
discrete alarms
   1: '', class Errors, trigger "Alarm0Pack16B_Alarmas_word" bit 0
   2: '', class Errors, trigger "Alarm0Pack16B_Alarmas_word" bit 1
   3: '', class Errors, trigger "Alarm0Pack16B_Alarmas_word" bit 2
   4: '', class Errors, trigger "Alarm0Pack16B_Alarmas_word" bit 3
   5: '', class Errors, trigger "Alarm0Pack16B_Alarmas_word" bit 4
   6: '', class Errors, trigger "Alarm0Pack16B_Alarmas_word" bit 5
   7: '', class Errors, trigger "Alarm0Pack16B_Alarmas_word" bit 6
   8: '', class Errors, trigger "Alarm0Pack16B_Alarmas_word" bit 7
   9: '', class Errors, trigger "Alarm0Pack16B_Alarmas_word" bit 8
   10: '', class Errors, trigger "Alarm0Pack16B_Alarmas_word" bit 9
   11: '', class Errors, trigger "Alarm0Pack16B_Alarmas_word" bit 10
   12: '', class Errors, trigger "Alarm0Pack16B_Alarmas_word" bit 11
   13: '', class Errors, trigger "Alarm0Pack16B_Alarmas_word" bit 12
   14: '', class Errors, trigger "Alarm0Pack16B_Alarmas_word" bit 13
   15: '', class Errors, trigger "Alarm0Pack16B_Alarmas_word" bit 14
   16: '', class Errors, trigger "Alarm0Pack16B_Alarmas_word" bit 15
   17: 'PeakDisplayPreAlarmHI', class Errors, trigger "Alarm1Pack16B_Alarmas_word" bit 0
   18: 'PeakDisplayAlarmHI', class Errors, trigger "Alarm1Pack16B_Alarmas_word" bit 1
   19: 'PeakDisplayPreAlarmLOW', class Errors, trigger "Alarm1Pack16B_Alarmas_word" bit 2
   20: 'PeakDisplayAlarmLOW', class Errors, trigger "Alarm1Pack16B_Alarmas_word" bit 3
   21: 'PlateauDisplayPreAlarmHI', class Errors, trigger "Alarm1Pack16B_Alarmas_word" bit 4
   22: 'PlateauDisplayAlarmHI', class Errors, trigger "Alarm1Pack16B_Alarmas_word" bit 5
   23: 'PlateauDisplayPreAlarmLOW', class Errors, trigger "Alarm1Pack16B_Alarmas_word" bit 6
   24: 'PlateaukDisplayAlarmLOW', class Errors, trigger "Alarm1Pack16B_Alarmas_word" bit 7
   25: 'PeepDisplayPreAlarmHI', class Errors, trigger "Alarm1Pack16B_Alarmas_word" bit 8
   26: 'PeepDisplayAlarmHI', class Errors, trigger "Alarm1Pack16B_Alarmas_word" bit 9
   27: 'PeepDisplayPreAlarmLOW', class Errors, trigger "Alarm1Pack16B_Alarmas_word" bit 10
   28: 'PeepDisplayAlarmLOW', class Errors, trigger "Alarm1Pack16B_Alarmas_word" bit 11
   29: 'FrequenciaDisplayPreAlarm / FrequencyDisplayPreAlarm', class Errors, trigger "Alarm1Pack16B_Alarmas_word" bit 12
   30: 'FrequenciaDisplayAlarmHI / FrequencyDisplayAlarmHI', class Errors, trigger "Alarm1Pack16B_Alarmas_word" bit 13
   31: 'FrequenciaDisplayPreAlarmLOW / FrequencyDisplayPreAlarmLOW', class Errors, trigger "Alarm1Pack16B_Alarmas_word" bit 14
   32: 'FrequenciaDisplayAlarmLOW / FrequencyDisplayAlarmLOW', class Errors, trigger "Alarm1Pack16B_Alarmas_word" bit 15
   33: 'TidalVolumeDisplayPreAlarm', class Errors, trigger "Alarm2Pack16B_Alarmas_word" bit 0
   34: 'TidalVolumeDisplayAlarmHI', class Errors, trigger "Alarm2Pack16B_Alarmas_word" bit 1
   35: 'TidalVolumeDisplayPreAlarmLOW', class Errors, trigger "Alarm2Pack16B_Alarmas_word" bit 2
   36: 'TidalVolumeDisplayAlarmLOW', class Errors, trigger "Alarm2Pack16B_Alarmas_word" bit 3
   37: 'MinuteVolumeDisplayPreAlarm', class Errors, trigger "Alarm2Pack16B_Alarmas_word" bit 4
   38: 'MinuteVolumeDisplayAlarmHI', class Errors, trigger "Alarm2Pack16B_Alarmas_word" bit 5
   39: 'MinuteVolumeDisplayPreAlarmLOW', class Errors, trigger "Alarm2Pack16B_Alarmas_word" bit 6
   40: 'MinuteVolumeDisplayAlarmLOW', class Errors, trigger "Alarm2Pack16B_Alarmas_word" bit 7
   41: 'TriggerDisplayPreAlarm', class Errors, trigger "Alarm2Pack16B_Alarmas_word" bit 8
   42: 'TriggerVolumeDisplayAlarmHI', class Errors, trigger "Alarm2Pack16B_Alarmas_word" bit 9
   43: 'TriggerVolumeDisplayPreAlarmLOW', class Errors, trigger "Alarm2Pack16B_Alarmas_word" bit 10
   44: 'TriggerVolumeDisplayAlarmLOW', class Errors, trigger "Alarm2Pack16B_Alarmas_word" bit 11
   45: 'BatteryDisplayPreAlarmHI', class Errors, trigger "Alarm2Pack16B_Alarmas_word" bit 12
   46: 'BatteryDisplayAlarmHI', class Errors, trigger "Alarm2Pack16B_Alarmas_word" bit 13
   47: 'BatteryDisplayPreAlarmLOW', class Errors, trigger "Alarm2Pack16B_Alarmas_word" bit 14
   48: 'BatteryDisplayAlarmLOW', class Errors, trigger "Alarm2Pack16B_Alarmas_word" bit 15
   49: '', class Errors, trigger "Alarm3Pack16B_Alarmas_word" bit 0
   50: '', class Errors, trigger "Alarm3Pack16B_Alarmas_word" bit 1
   51: '', class Errors, trigger "Alarm3Pack16B_Alarmas_word" bit 2
   52: '', class Errors, trigger "Alarm3Pack16B_Alarmas_word" bit 3
   53: '', class Errors, trigger "Alarm3Pack16B_Alarmas_word" bit 4
   54: '', class Errors, trigger "Alarm3Pack16B_Alarmas_word" bit 5
   55: '', class Errors, trigger "Alarm3Pack16B_Alarmas_word" bit 6
   56: '', class Errors, trigger "Alarm3Pack16B_Alarmas_word" bit 7
   57: '', class Errors, trigger "Alarm3Pack16B_Alarmas_word" bit 8
   58: '', class Errors, trigger "Alarm3Pack16B_Alarmas_word" bit 9
   59: '', class Errors, trigger "Alarm3Pack16B_Alarmas_word" bit 10
   60: '', class Errors, trigger "Alarm3Pack16B_Alarmas_word" bit 11
   61: '', class Errors, trigger "Alarm3Pack16B_Alarmas_word" bit 12
   62: '', class Errors, trigger "Alarm3Pack16B_Alarmas_word" bit 13
   63: '', class Errors, trigger "Alarm3Pack16B_Alarmas_word" bit 14
   64: '', class Errors, trigger "Alarm3Pack16B_Alarmas_word" bit 15

text list "PatientSex": 1 'Man'; 2 'Mujer / Woman'; 0 'No Seleccionado / Not Selected'

text list "ControlMode": 0 'NO SELECCIONADO / NOT SELECTED'; 1 'CP Control Presión / PC Pressure Control'; 2 'CV Control Volumen / VC Volume Control'; 3 'CC Control Caudal / FC Flow Control'

text list "ModeSelected": 0 'Modo NS / NC Mode'; 1 'Modo CP / PC Mode'; 2 'CV Modo / VC Mode'; 3 'CF Modo / FC Mode'

screen "Start" 800x480
   GraphicView "Visor de gráficos_1" at 8,10 size 785x426; Picture "covid19"
   TextField "Campo de texto_1" at 30,81 size 657x91; Text 'Reespirator-2020'
   IOField "Campo ES_1" at 593,393 size 191x32; FormatPattern 9999999999999999999999999999999999999999
      ProcessValue <- "DateTime_LocalDateOut"
   TextField "Campo de texto_2" at 90,188 size 363x62; Text 'De personas, / From people, / From persons,'
   TextField "Campo de texto_3" at 290,250 size 405x62; Text 'para PERSONAS / for PEOPLE'
   Button "Botón_1" at 7,442 size 80x35; TextOff 'GRAFICOS / GRAPHICS'
      on Press: ActivateScreen("Graphics", 0)
   Button "Botón_3" at 92,442 size 80x35; TextOff 'DATOS / DATA'
      on Press: ActivateScreen("Parameters", 0)
   Button "Botón_4" at 347,442 size 80x35; TextOff 'MANUALES / MANUALS'
      on Press: ActivateScreen("UserManual", 0)
   Button "Botón_5" at 432,442 size 80x35; TextOff 'ALARMAS / ALARMS'
      on Press: ActivateScreen("Alarms", 0)
   Button "Botón_6" at 177,442 size 80x35; TextOff 'PACIENTE / PATIENT'
      on Press: function_efd93a16("PatientData", 0, 0, 1, -1, 1)
   TextField "Campo de texto_9" at 526,445 size 101x27; Text 'BATERIA / BATTERY'
   IOField "Campo ES_14" at 621,442 size 89x35; FormatPattern 99.9; Unit  Vdc
      ProcessValue <- "DataValues_BatteryVoltage"
   Button "Botón_11" at 534,442 size 35x35; TextOff 'M'
      on Press: ActivateScreen("Start", 0)
   IOField "Campo ES_15" at 713,442 size 82x35; FormatPattern 999.9; Unit  %
      ProcessValue <- "DataValues_BatteryCapacity"
   Button "Botón_8" at 582,442 size 35x35; TextOff 'M'
      on Press: ActivateScreen("Motor", 0)
   Button "Botón_2" at 262,442 size 80x35; TextOff 'RPM / BPM'
      on Press: function_efd93a16("RespirationRatios", 0, 0, 1, -1, 1)
   Button "Botón_7" at 20,366 size 100x60; TextOff 'Text'; PictureOff "spain_flags_flag_17068"
      on Click: function_fb9197e8(L es-ES)
   Button "Botón_10" at 124,367 size 100x60; TextOff 'Text'; PictureOff "united_kingdom_flags_flag_17079"
      on Click: function_fb9197e8(L en-GB)
   Button "Botón_9" at 228,367 size 100x60; TextOff 'Text'; PictureOff "france_flags_flag_16999"
      on Click: function_fb9197e8(L fr-FR)
   Button "Botón_12" at 332,368 size 100x60; TextOff 'Text'; PictureOff "portugal_flags_flag_17054"
      on Click: function_fb9197e8(L pt-PT)

screen "Parameters" 800x480
   TextField "Campo de texto_3" at 181,181 size 19x29; Text 'Text'
   IOField "Campo ES_8" at 352,69 size 75x35; Authorization "Operación"; FormatPattern 999
      ProcessValue <- "DataValues_PipValue"
   IOField "Campo ES_2" at 256,69 size 75x35; FormatPattern 999
      ProcessValue <- "OperatingParameters_PipMax"
   IOField "Campo ES_3" at 15,69 size 75x35; FormatPattern 999
      ProcessValue <- "OperatingParameters_PipSetpoint"
      Visibility <- "OperatingParameters_ControlMode"
   IOField "Campo ES_4" at 352,123 size 75x35; Authorization "Operación"; FormatPattern 999
      ProcessValue <- "DataValues_PlateauValue"
   IOField "Campo ES_6" at 256,123 size 75x35; FormatPattern 999
      ProcessValue <- "OperatingParameters_PlateauMax"
   IOField "Campo ES_9" at 352,178 size 75x35; FormatPattern 999
      ProcessValue <- "DataValues_PeepValue"
   IOField "Campo ES_11" at 256,178 size 75x35; FormatPattern 999
      ProcessValue <- "OperatingParameters_PeepMax"
   IOField "Campo ES_12" at 15,178 size 75x35; FormatPattern 999
      ProcessValue <- "OperatingParameters_PeepSetpoint"
   IOField "Campo ES_13" at 352,232 size 75x35; FormatPattern 999
      ProcessValue <- "DataValues_FrequencyValue"
   IOField "Campo ES_17" at 256,232 size 75x35; FormatPattern 999
      ProcessValue <- "OperatingParameters_FrequencyMax"
   IOField "Campo ES_18" at 15,232 size 75x35; FormatPattern 999
      ProcessValue <- "OperatingParameters_FrequencySetpoint"
   IOField "Campo ES_19" at 352,286 size 75x35; FormatPattern 999
      ProcessValue <- "DataValues_TidalVolumeValue"
   IOField "Campo ES_21" at 256,286 size 75x35; FormatPattern 999
      ProcessValue <- "OperatingParameters_TidalVolumenMax"
   IOField "Campo ES_23" at 352,340 size 75x35; FormatPattern 999
      ProcessValue <- "DataValues_MinumValue"
   IOField "Campo ES_25" at 256,340 size 75x35; FormatPattern 999
      ProcessValue <- "OperatingParameters_MinimumVolumeMax"
   IOField "Campo ES_29" at 14,394 size 75x35; FormatPattern 999
      ProcessValue <- "OperatingParameters_TriggerSetpoint"
   TextField "Campo de texto_6" at 266,18 size 55x29; Text 'MAX'
   TextField "Campo de texto_7" at 351,18 size 81x29; Text 'VALOR / VALUE'
   TextField "Campo de texto_8" at 460,18 size 56x29; Text 'MIN'
   TrendView "Visor de curvas_2" at 533,145 size 255x294
   TrendView "Visor de curvas_1" at 533,8 size 254x137
   IOField "Campo ES_7" at 449,69 size 75x35; FormatPattern 999
      ProcessValue <- "OperatingParameters_PipMin"
   IOField "Campo ES_22" at 450,123 size 75x35; FormatPattern 999
      ProcessValue <- "OperatingParameters_PlateauMin"
   IOField "Campo ES_26" at 450,178 size 75x35; FormatPattern 999
      ProcessValue <- "OperatingParameters_PeepMin"
   IOField "Campo ES_27" at 449,232 size 75x35; FormatPattern 999
      ProcessValue <- "OperatingParameters_FrequencyMin"
   IOField "Campo ES_28" at 450,286 size 75x35; FormatPattern 999
      ProcessValue <- "OperatingParameters_TidalVolumenMin"
   IOField "Campo ES_30" at 450,340 size 75x35; FormatPattern 999
      ProcessValue <- "OperatingParameters_MinimumVolumeMin"
   Button "Botón_7" at 92,394 size 53x35; TextOff 'Trigger'
      Visibility <- "Clock_1Hz"
   IOField "Campo ES_1" at 15,17 size 242x32; FormatPattern 99999999999999999999
      ProcessValue <- "DateTime_LocalDateOut"
   GraphicIOField "PlotLight_Round_GN" at 333,69 size 17x17; PictureOff "gris"; PictureOn "rojo"
      ProcessValue <- "AlarmsRaw_PipDisplayAlarmHI"
   GraphicIOField "PlotLight_Round_GN_1" at 333,123 size 17x17; PictureOff "gris"; PictureOn "rojo"
      ProcessValue <- "AlarmsRaw_PlateauDisplayAlarmHI"
   GraphicIOField "PlotLight_Round_GN_2" at 333,178 size 17x17; PictureOff "gris"; PictureOn "rojo"
      ProcessValue <- "AlarmsRaw_PeepDisplayAlarmHI"
   GraphicIOField "PlotLight_Round_GN_3" at 333,232 size 17x17; PictureOff "gris"; PictureOn "rojo"
      ProcessValue <- "AlarmsRaw_FrequencyDisplayAlarmHI"
   GraphicIOField "PlotLight_Round_GN_4" at 333,286 size 17x17; PictureOff "gris"; PictureOn "rojo"
      ProcessValue <- "AlarmsRaw_TidalVolumeDisplayAlarmHI"
   GraphicIOField "PlotLight_Round_GN_5" at 333,340 size 17x17; PictureOff "gris"; PictureOn "rojo"
      ProcessValue <- "AlarmsRaw_VolumeMinuteDisplayAlarmHI"
   GraphicIOField "PlotLight_Round_GN_6" at 430,87 size 17x17; PictureOn "rojo"; PictureOff "gris"
      ProcessValue <- "AlarmsRaw_PipDisplayAlarmLOW"
   GraphicIOField "PlotLight_Round_GN_7" at 430,141 size 17x17; PictureOn "rojo"; PictureOff "gris"
      ProcessValue <- "AlarmsRaw_PlateauDisplayAlarmLOW"
   GraphicIOField "PlotLight_Round_GN_8" at 430,196 size 17x17; PictureOn "rojo"; PictureOff "gris"
      ProcessValue <- "AlarmsRaw_PeepDisplayAlarmLOW"
   GraphicIOField "PlotLight_Round_GN_9" at 430,250 size 17x17; PictureOn "rojo"; PictureOff "gris"
      ProcessValue <- "AlarmsRaw_FrequencyDisplayAlarmLOW"
   GraphicIOField "PlotLight_Round_GN_10" at 430,304 size 17x17; PictureOn "rojo"; PictureOff "gris"
      ProcessValue <- "AlarmsRaw_TidalVolumeDisplayAlarmLOW"
   GraphicIOField "PlotLight_Round_GN_11" at 430,358 size 17x17; PictureOn "rojo"; PictureOff "gris"
      ProcessValue <- "AlarmsRaw_VolumeMinuteDisplayAlarmLOW"
   GraphicIOField "PlotLight_Round_GN_12" at 333,87 size 17x17; PictureOff "gris"; PictureOn "amarillo"
      ProcessValue <- "AlarmsRaw_PipDisplayPreAlarmHI"
   GraphicIOField "PlotLight_Round_GN_13" at 333,141 size 17x17; PictureOff "gris"; PictureOn "amarillo"
      ProcessValue <- "AlarmsRaw_PlateauDisplayPreAlarmHI"
   GraphicIOField "PlotLight_Round_GN_14" at 333,196 size 17x17; PictureOff "gris"; PictureOn "amarillo"
      ProcessValue <- "AlarmsRaw_PeepDisplayPreAlarmHI"
   GraphicIOField "PlotLight_Round_GN_15" at 333,250 size 17x17; PictureOff "gris"; PictureOn "amarillo"
      ProcessValue <- "AlarmsRaw_FrequencyDisplayPreAlarmHI"
   GraphicIOField "PlotLight_Round_GN_16" at 333,304 size 17x17; PictureOff "gris"; PictureOn "amarillo"
      ProcessValue <- "AlarmsRaw_TidalVolumeDisplayPreAlarmHI"
   GraphicIOField "PlotLight_Round_GN_17" at 333,358 size 17x17; PictureOff "gris"; PictureOn "amarillo"
      ProcessValue <- "AlarmsRaw_VolumeMinuteDisplayPreAlarmHI"
   GraphicIOField "PlotLight_Round_GN_18" at 430,69 size 17x17; PictureOn "amarillo"; PictureOff "gris"
      ProcessValue <- "AlarmsRaw_PipDisplayPreAlarmLOW"
   GraphicIOField "PlotLight_Round_GN_19" at 430,123 size 17x17; PictureOn "amarillo"; PictureOff "gris"
      ProcessValue <- "AlarmsRaw_PlateauDisplayPreAlarmLOW"
   GraphicIOField "PlotLight_Round_GN_20" at 430,178 size 17x17; PictureOn "amarillo"; PictureOff "gris"
      ProcessValue <- "AlarmsRaw_PeepDisplayPreAlarmLOW"
   GraphicIOField "PlotLight_Round_GN_21" at 430,232 size 17x17; PictureOn "amarillo"; PictureOff "gris"
      ProcessValue <- "AlarmsRaw_FrequencyDisplayPreAlarmLOW"
   GraphicIOField "PlotLight_Round_GN_22" at 430,286 size 17x17; PictureOn "amarillo"; PictureOff "gris"
      ProcessValue <- "AlarmsRaw_TidalVolumeDisplayPreAlarmLOW"
   GraphicIOField "PlotLight_Round_GN_23" at 430,340 size 17x17; PictureOn "amarillo"; PictureOff "gris"
      ProcessValue <- "AlarmsRaw_VolumeMinuteDisplayPreAlarmLOW"
   Button "Botón_9" at 100,69 size 144x35; TextOff 'PIP'
      on Press: function_efd93a16("Pip", 0, 0, -1, -1, 1)
   Button "Botón_10" at 102,123 size 144x35; TextOff 'PLATEAU'
      on Press: function_efd93a16("Plateau", 0, 0, -1, -1, 1)
   Button "Botón_12" at 101,178 size 144x35; TextOff 'PEEP'
      on Press: function_efd93a16("Peep", 0, 0, -1, -1, 1)
   Button "Botón_13" at 102,232 size 144x35; TextOff 'FRECUENCIA / FREQUENCY'
      on Press: function_efd93a16("Frecuency", 0, 0, -1, -1, 1)
   Button "Botón_14" at 100,286 size 144x35; TextOff 'VOL TIDAL / TIDAL VOL'
      on Press: function_efd93a16("TidalVolume", 0, 0, -1, -1, 1)
   Button "Botón_15" at 100,340 size 144x35; TextOff 'VOL. MINUTO / VOL. MINUTE'
      on Press: function_efd93a16("VolumeMinute", 0, 0, -1, -1, 1)
   Button "Botón_16" at 149,395 size 135x35; TextOff 'TRIGGER'
      on Press: function_efd93a16("Trigger", 0, 0, -1, -1, 1)
   TextField "Campo de texto_2" at 289,395 size 61x35; Text 'OFF'
      Visibility <- "OperatingParameters_Trigger"
   TextField "Campo de texto_10" at 289,395 size 61x35; Text 'ON'
      Visibility <- "OperatingParameters_Trigger"
   Button "Botón_2" at 289,395 size 61x35; TextOn 'ON'; TextOff 'Text'
      on Click: InvertBit("OperatingParameters_Trigger")
      Appearance <- "OperatingParameters_Trigger"
   Button "Botón_17" at 372,396 size 150x35; TextOff 'ENTORNO / ENVIROMENT'
      on Press: function_efd93a16("Enviroment", 0, 0, -1, -1, 1)
   TextField "Campo de texto_9" at 526,445 size 101x27; Text 'BATERIA / BATTERY'
   IOField "Campo ES_14" at 621,442 size 89x35; FormatPattern 99.9; Unit  Vdc
      ProcessValue <- "DataValues_BatteryVoltage"
   Button "Botón_11" at 534,442 size 35x35; TextOff 'M'
      on Press: ActivateScreen("Start", 0)
   IOField "Campo ES_15" at 713,442 size 82x35; FormatPattern 999.9; Unit  %
      ProcessValue <- "DataValues_BatteryCapacity"
   Button "Botón_8" at 582,442 size 35x35; TextOff 'M'
      on Press: ActivateScreen("Motor", 0)
   IOField "Campo ES_10" at 15,286 size 75x35; FormatPattern 999
      ProcessValue <- "OperatingParameters_TidalVolumenSetpoint"
      Visibility <- "OperatingParameters_ControlMode"
   IOField "Campo ES_16" at 15,340 size 75x35; FormatPattern 999
      ProcessValue <- "OperatingParameters_MinimumVolumeSetpoint"
      Visibility <- "OperatingParameters_ControlMode"
   Button "Botón_1" at 7,442 size 80x35; TextOff 'GRAFICOS / GRAPHICS'
      on Press: ActivateScreen("Graphics", 0)
   Button "Botón_3" at 92,442 size 80x35; TextOff 'DATOS / DATA'
      on Press: ActivateScreen("Parameters", 0)
   Button "Botón_4" at 347,442 size 80x35; TextOff 'MANUALES / MANUALS'
      on Press: ActivateScreen("UserManual", 0)
   Button "Botón_5" at 432,442 size 80x35; TextOff 'ALARMAS / ALARMS'
      on Press: ActivateScreen("Alarms", 0)
   Button "Botón_6" at 177,442 size 80x35; TextOff 'PACIENTE / PATIENT'
      on Press: function_efd93a16("PatientData", 0, 0, 1, -1, 1)
   Button "Botón_18" at 262,442 size 80x35; TextOff 'RPM / BPM'
      on Press: function_efd93a16("RespirationRatios", 0, 0, 1, -1, 1)
   Button "Botón_19" at 7,2 size 35x28; TextOff 'M'
      on Press: ActivateScreen("Start", 0)
   Button "Botón_20" at 86,2 size 35x29; TextOff 'M'
      on Press: ActivateScreen("Motor", 0)

screen "UserManual" 800x480
   PDFView "Visor de PDF_1" at 0,1 size 800x437
   TextField "Campo de texto_9" at 526,445 size 101x27; Text 'BATERIA / BATTERY'
   IOField "Campo ES_14" at 621,442 size 89x35; FormatPattern 99.9; Unit  Vdc
      ProcessValue <- "DataValues_BatteryVoltage"
   Button "Botón_11" at 534,442 size 35x35; TextOff 'M'
      on Press: ActivateScreen("Start", 0)
   IOField "Campo ES_15" at 713,442 size 82x35; FormatPattern 999.9; Unit  %
      ProcessValue <- "DataValues_BatteryCapacity"
   Button "Botón_8" at 582,442 size 35x35; TextOff 'M'
      on Press: ActivateScreen("Motor", 0)
   Button "Botón_1" at 7,442 size 80x35; TextOff 'GRAFICOS / GRAPHICS'
      on Press: ActivateScreen("Graphics", 0)
   Button "Botón_3" at 92,442 size 80x35; TextOff 'DATOS / DATA'
      on Press: ActivateScreen("Parameters", 0)
   Button "Botón_4" at 347,442 size 80x35; TextOff 'MANUALES / MANUALS'
      on Press: ActivateScreen("UserManual", 0)
   Button "Botón_5" at 432,442 size 80x35; TextOff 'ALARMAS / ALARMS'
      on Press: ActivateScreen("Alarms", 0)
   Button "Botón_6" at 177,442 size 80x35; TextOff 'PACIENTE / PATIENT'
      on Press: function_efd93a16("PatientData", 0, 0, 1, -1, 1)
   Button "Botón_2" at 262,442 size 80x35; TextOff 'RPM / BPM'
      on Press: function_efd93a16("RespirationRatios", 0, 0, 1, -1, 1)

screen "Alarms" 800x480
   AlarmView "Visor de avisos_1" at 0,35 size 799x403
      Visibility <- "AlwaysTRUE"
   IOField "Campo ES_1" at 607,2 size 191x32; FormatPattern 9999999999999999999999999999999999999999
      ProcessValue <- "DateTime_LocalDateOut"
   TextField "Campo de texto_1" at 0,6 size 204x29; Text 'Reespirator-2020'
   TextField "Campo de texto_2" at 318,5 size 113x29; Text 'ALARMAS / ALARMS'
   TextField "Campo de texto_9" at 526,445 size 101x27; Text 'BATERIA / BATTERY'
   IOField "Campo ES_14" at 621,442 size 89x35; FormatPattern 99.9; Unit  Vdc
      ProcessValue <- "DataValues_BatteryVoltage"
   IOField "Campo ES_15" at 713,442 size 82x35; FormatPattern 999.9; Unit  %
      ProcessValue <- "DataValues_BatteryCapacity"
   Button "Botón_1" at 7,442 size 80x35; TextOff 'GRAFICOS / GRAPHICS'
      on Press: ActivateScreen("Graphics", 0)
   Button "Botón_3" at 92,442 size 80x35; TextOff 'DATOS / DATA'
      on Press: ActivateScreen("Parameters", 0)
   Button "Botón_4" at 347,442 size 80x35; TextOff 'MANUALES / MANUALS'
      on Press: ActivateScreen("UserManual", 0)
   Button "Botón_5" at 432,442 size 80x35; TextOff 'ALARMAS / ALARMS'
      on Press: ActivateScreen("Alarms", 0)
   Button "Botón_6" at 177,442 size 80x35; TextOff 'PACIENTE / PATIENT'
      on Press: function_efd93a16("PatientData", 0, 0, 1, -1, 1)
   Button "Botón_2" at 262,442 size 80x35; TextOff 'RPM / BPM'
      on Press: function_efd93a16("RespirationRatios", 0, 0, 1, -1, 1)
   Button "Botón_16" at 7,2 size 35x28; TextOff 'M'
      on Press: ActivateScreen("Start", 0)
   Button "Botón_17" at 86,2 size 35x29; TextOff 'M'
      on Press: ActivateScreen("Motor", 0)
   Button "Botón_11" at 534,442 size 35x35; TextOff 'M'
      on Press: ActivateScreen("Start", 0)
   Button "Botón_8" at 582,442 size 35x35; TextOff 'M'
      on Press: ActivateScreen("Motor", 0)

screen "Motor" 800x480
   Button "Botón_2" at 73,9 size 145x40; TextOn 'Habilitado / ENABLED'; TextOff 'HABILITACION POTENCIA / POWER ENABLE'
      on Press: InvertBit("MotorControl_POWER_Enable")
   Button "Botón_6" at 73,57 size 145x40; TextOff 'RESET'
      on Press: function_b14e0dd5("MotorControl_RESET_Execute", 0)
   Button "Botón_7" at 73,118 size 145x40; TextOff 'RETORNO / HOME'
      on Press: function_b14e0dd5("MotorControl_HOME_Execute", 0)
   Button "Botón_8" at 295,9 size 145x40; TextOff 'Paro / HALT'
      on Press: function_b14e0dd5("MotorControl_HALT_Execute", 0)
   IOField "Campo ES_2" at 522,312 size 145x40; FormatPattern 9999
      ProcessValue <- "MotorControl_ABSOLUTE_Velocity"
   IOField "Campo ES_6" at 244,118 size 142x40; FormatPattern 9999
      ProcessValue <- "MotorControl_HOME_Position"
   Button "Botón_11" at 73,312 size 145x40; TextOff 'ABS EXECUTE'
      on Press: function_b14e0dd5("MotorControl_ABSOLUTE_Execute", 0)
   Button "Botón_13" at 610,117 size 145x40; TextOff 'HABILITACION PWM / PWM ENABLE'
      on Press: InvertBit("2_PWMValve_Enable")
   Rectangle "Rectángulo_5" at 259,8 size 15x41
      Visibility <- "MotorControl_HALT_Execute"
   Rectangle "Rectángulo_11" at 275,8 size 15x41
      Visibility <- "MotorControl_HALT_Error"
   Rectangle "Rectángulo_12" at 243,8 size 15x41
      Visibility <- "MotorControl_HALT_Done"
   Rectangle "Rectángulo_3" at 34,9 size 15x41
      Visibility <- "MotorControl_POWER_Enable"
   Rectangle "Rectángulo_4" at 50,9 size 15x41
      Visibility <- "MotorControl_POWER_Error"
   Rectangle "Rectángulo_6" at 18,9 size 15x41
      Visibility <- "MotorControl_POWER_Status"
   Rectangle "Rectángulo_7" at 35,56 size 15x41
      Visibility <- "MotorControl_RESET_Execute"
   Rectangle "Rectángulo_10" at 51,56 size 15x41
      Visibility <- "MotorControl_RESET_Error"
   Rectangle "Rectángulo_13" at 19,56 size 15x41
      Visibility <- "MotorControl_RESET_Done"
   Rectangle "Rectángulo_14" at 36,118 size 15x41
      Visibility <- "MotorControl_HOME_Execute"
   Rectangle "Rectángulo_15" at 52,118 size 15x41
      Visibility <- "MotorControl_HOME_Error"
   Rectangle "Rectángulo_16" at 20,118 size 15x41
      Visibility <- "MotorControl_HOME_Done"
   IOField "Campo ES_5" at 244,312 size 145x40; FormatPattern 9999
      ProcessValue <- "MotorControl_ABSOLUTE_Position"
   Rectangle "Rectángulo_24" at 36,312 size 15x41
      Visibility <- "MotorControl_ABSOLUTE_Execute"
   Rectangle "Rectángulo_25" at 52,312 size 15x41
      Visibility <- "MotorControl_ABSOLUTE_Error"
   Rectangle "Rectángulo_26" at 20,312 size 15x41
      Visibility <- "MotorControl_ABSOLUTE_Done"
   IOField "Campo ES_1" at 522,377 size 145x40; FormatPattern 9999
      ProcessValue <- "MotorControl_RELATIVE_Velocity"
   Button "Botón_15" at 73,377 size 145x40; TextOff 'REL EXECUTE'
      on Press: function_b14e0dd5("MotorControl_RELATIVE_Execute", 0)
   IOField "Campo ES_4" at 244,377 size 145x40; FormatPattern 9999
      ProcessValue <- "MotorControl_RELATIVE_Distance"
   Rectangle "Rectángulo_28" at 36,377 size 15x41
      Visibility <- "MotorControl_RELATIVE_Execute"
   Rectangle "Rectángulo_29" at 52,377 size 15x41
      Visibility <- "MotorControl_RELATIVE_Error"
   Rectangle "Rectángulo_30" at 20,377 size 15x41
      Visibility <- "MotorControl_RELATIVE_Done"
   TextField "Campo de texto_4" at 394,318 size 100x29; Text 'Posición / Position'
   TextField "Campo de texto_6" at 394,382 size 104x29; Text 'Distance'
   TextField "Campo de texto_7" at 676,318 size 115x29; Text 'Velocidad / Velocity'
   TextField "Campo de texto_8" at 676,382 size 115x29; Text 'Velocidad / Velocity'
   Button "Botón_16" at 609,249 size 145x40; TextOff 'JOG FORWARD'
      on Press: function_b14e0dd5("MotorControl_JOG_Forward", 0)
   Button "Botón_17" at 73,247 size 145x40; TextOff 'JOG BACKWARD'
      on Press: function_b14e0dd5("MotorControl_JOG_Backward", 0)
   IOField "Campo ES_3" at 245,248 size 145x40; FormatPattern 9999
      ProcessValue <- "MotorControl_JOG_Velocity"
   Rectangle "Rectángulo_32" at 573,248 size 15x41
      Visibility <- "MotorControl_JOG_Forward"
   Rectangle "Rectángulo_33" at 589,248 size 15x41
      Visibility <- "MotorControl_JOG_Error"
   Rectangle "Rectángulo_34" at 557,248 size 15x41
      Visibility <- "MotorControl_JOG_Invelocity"
   Rectangle "Rectángulo_35" at 37,246 size 15x41
      Visibility <- "MotorControl_JOG_Backward"
   Rectangle "Rectángulo_36" at 53,246 size 15x41
      Visibility <- "MotorControl_JOG_Error"
   Rectangle "Rectángulo_37" at 21,246 size 15x41
      Visibility <- "MotorControl_JOG_Invelocity"
   TextField "Campo de texto_2" at 397,253 size 115x29; Text 'Velocidad / Velocity'
   TextField "Campo de texto_3" at 397,123 size 100x29; Text 'Posición / Position'
   Button "Botón_10" at 71,183 size 145x40; TextOff 'VELOCIDAD / VELOCITY'
      on Press: function_b14e0dd5("MotorControl_Velocity_Execute", 0)
   IOField "Campo ES_29" at 243,184 size 145x40; FormatPattern 9999